// TIA Portal project "Catalyst_syzygy_v2.1" (V17)

(* hardware
DEVICE "S7-1500R/H system_1"  S7-1500R/H-Station
   slot 0: "Rail_0"  Rack  6ES7 590-1***0-0AA0
   slot 1: "Rail_1"  Rack  6ES7 590-1***0-0AA0
   slot 1: "Catalyst_PLC_1"  CPU 1515R-2 PN  6ES7 515-2RM00-0AB0  V2.9
      slot 3: "CPU display_1"  6ES7591-1BA00-0AA0
      slot 32768: "PROFINET interface_1"  X1
         slot 32769: "Port_1"  X1 P1
         slot 32770: "Port_2"  X1 P2
      slot 33024: "PROFINET interface_2"  X2
         slot 33025: "Port_1"  X2 P1
   slot 1: "Catalyst_PLC_2"  CPU 1515R-2 PN  6ES7 515-2RM00-0AB0  V2.9
      slot 3: "CPU display_1"  6ES7591-1BA00-0AA0
      slot 32768: "PROFINET interface_1"  X1
         slot 32769: "Port_1"  X1 P1
         slot 32770: "Port_2"  X1 P2
      slot 33024: "PROFINET interface_2"  X2
         slot 33025: "Port_1"  X2 P1
DEVICE "S7-1500/ET200MP station_1"  S7-1500 station
   slot 0: "Rail_0"  Rack  6ES7 590-1***0-0AA0
   slot 1: "CatalystLocalIO_02"  IM 155-5 PN HF  6ES7 155-5AA00-0AC0  V4.2
   slot 2: "LocalIO_02_AI_01"  AI 8xU/I/RTD/TC ST  6ES7 531-7KF00-0AB0  V2.2
   slot 3: "LocalIO_02_AI_02"  AI 8xU/I/RTD/TC ST  6ES7 531-7KF00-0AB0  V2.2
   slot 4: "LocalIO_02_AI_03"  AI 8xU/I/RTD/TC ST  6ES7 531-7KF00-0AB0  V2.2
   slot 5: "LocalIO_02_AI_04"  AI 8xU/I/RTD/TC ST  6ES7 531-7KF00-0AB0  V2.2
   slot 6: "LocalIO_02_AI_05"  AI 8xU/I/RTD/TC ST  6ES7 531-7KF00-0AB0  V2.2
   slot 7: "LocalIO_02_AI_06"  AI 8xU/I/RTD/TC ST  6ES7 531-7KF00-0AB0  V2.2
   slot 8: "LocalIO_02_AI_07"  AI 8xU/I/RTD/TC ST  6ES7 531-7KF00-0AB0  V2.2
   slot 9: "LocalIO_02_AQ_01"  AQ 8xU/I HS  6ES7 532-5HF00-0AB0  V2.2
   slot 10: "LocalIO_02_AQ_02"  AQ 8xU/I HS  6ES7 532-5HF00-0AB0  V2.1
   slot 11: "LocalIO_02_AQ_03"  AQ 8xU/I HS  6ES7 532-5HF00-0AB0  V2.2
DEVICE "S7-1500/ET200MP station_2"  S7-1500 station
   slot 0: "Rail_0"  Rack  6ES7 590-1***0-0AA0
   slot 1: "CatalystLocalIO_01"  IM 155-5 PN HF  6ES7 155-5AA00-0AC0  V4.4
   slot 2: "LocalIO_01_DI_01"  DI 16x24VDC HF  6ES7 521-1BH00-0AB0  V2.2
   slot 3: "LocalIO_01_DI_02"  DI 16x24VDC HF  6ES7 521-1BH00-0AB0  V2.2
   slot 4: "LocalIO_01_DI_03"  DI 16x24VDC HF  6ES7 521-1BH00-0AB0  V2.2
   slot 5: "LocalIO_01_DI_04"  DI 16x24VDC HF  6ES7 521-1BH00-0AB0  V2.2
   slot 6: "LocalIO_01_DI_05"  DI 16x24VDC HF  6ES7 521-1BH00-0AB0  V2.2
   slot 7: "LocalIO_01_DI_06"  DI 16x24VDC HF  6ES7 521-1BH00-0AB0  V2.2
   slot 8: "LocalIO_01_DQ_01"  DQ 16x24VDC/0.5A HF  6ES7 522-1BH01-0AB0  V1.1
   slot 9: "LocalIO_01_DQ_02"  DQ 16x24VDC/0.5A HF  6ES7 522-1BH01-0AB0  V1.1
   slot 10: "LocalIO_01_DQ_03"  DQ 16x24VDC/0.5A HF  6ES7 522-1BH01-0AB0  V1.1
   slot 11: "LocalIO_01_DQ_04"  DQ 16x24VDC/0.5A HF  6ES7 522-1BH01-0AB0  V1.1
   slot 12: "LocalIO_01_AI_01"  AI 8xU/I/RTD/TC ST  6ES7 531-7KF00-0AB0  V2.2
   slot 13: "LocalIO_01_AI_02"  AI 8xU/I/RTD/TC ST  6ES7 531-7KF00-0AB0  V2.2
   slot 14: "LocalIO_01_AI_03"  AI 8xU/I/RTD/TC ST  6ES7 531-7KF00-0AB0  V2.2
DEVICE "SITOP station_1"  SITOP-Station
   slot 0: "Rack_0"  Rail
   slot 0: "UPS1600"  UPS1600 40A PN  6EP4137-3AB00-2AY0  V2.5
   slot 1: "BAT1600 EX Pb 24V 12Ah_1"  Battery module EX 12Ah Pb  6EP4135-0GL00-0AY0  V1.0
DEVICE "GSD device_1"  GSD.Device.PN
   slot 0: "Rack"  Rack  V1.0
   slot 0: "R-402_DO"  FEN20-4DIP-4DXP  6931090  SW V 1.7.14
      slot 0: "DAP v3.1"  DAP v3.1
      slot 1: "PN-IO"  PN-IO
         slot 1: "Port 1"  Port 1
         slot 2: "Port 2"  Port 2
      slot 1: "4DIP-DXP_1"  4DIP-DXP
         slot 0: "4DIP-DXP"  4DIP-DXP
DEVICE "ET 200SP station_1"  ET 200SP-Station
   slot 0: "Rack_0"  Rack  6ES5 710-8MAx1
   slot 0: "Centrifuge_RIO"  IM 155-6 PN/2 HF  6ES7 155-6AU01-0CN0  V4.2
   slot 1: "DI 8x24VDC ST_1"  DI 8x24VDC ST  6ES7 131-6BF01-0BA0  V0.0
      slot 1: "DI 8x24VDC ST_1"  DI 8x24VDC ST
   slot 2: "DI 8x24VDC ST_2"  DI 8x24VDC ST  6ES7 131-6BF01-0BA0  V0.0
      slot 1: "DI 8x24VDC ST_2"  DI 8x24VDC ST
   slot 3: "DQ 8x24VDC/0.5A ST_1"  DQ 8x24VDC/0.5A ST  6ES7 132-6BF01-0BA0  V0.0
      slot 1: "DQ 8x24VDC/0.5A ST_1"  DQ 8x24VDC/0.5A ST
   slot 4: "AI 4xI 2-,4-wire ST_1"  AI 4xI 2-,4-wire ST  6ES7 134-6GD01-0BA1  V2.0
      slot 1: "AI 4xI 2-,4-wire ST_1"  AI 4xI 2-,4-wire ST
   slot 5: "AQ 4xU/I ST_1"  AQ 4xU/I ST  6ES7 135-6HD00-0BA1  V1.1
      slot 1: "AQ 4xU/I ST_1"  AQ 4xU/I ST
   slot 6: "Server module_1"  Server module  6ES7 193-6PA00-0AA0  V1.1
      slot 1: "Server module_1"  Server module
   slot 127: "BA 2xRJ45"  BA 2xRJ45  6ES7 193-6AR00-0AA0  V0.0
      slot 1: "Port_1"  X1 P1 R  6ES7 193-6AR00-0AA0  V0.0
      slot 2: "Port_2"  X1 P2 R  6ES7 193-6AR00-0AA0  V0.0
DEVICE "GSD device_2"  GSD.Device.PN
   slot 0: "Rack"  Rack  V1.0
   slot 0: "MIXER_T103_VFD"  SINAMICS G120C PN V4.7  6SL3 210-1KExx-xxFx  V4.70
      slot 0: "SINAMICS G120C PN V4.7"  SINAMICS G120C PN V4.7
      slot 1: "PN-IO"  PN-IO
         slot 1: "Port 1"  Port 1
         slot 2: "Port 2"  Port 2
      slot 1: "Drive_1"  Drive
         slot 0: "Module Access Point"  Module Access Point
   slot 2: "Standard telegram 1, PZD-2/2"  Standard telegram 1, PZD-2/2
*)

// ===== PLC "Catalyst_PLC_1"  CPU 1515R-2 PN =====

VAR_GLOBAL   // PLC tag table "Default tag table"
   "Tag_1" AT %T64435 : Timer;
   "Tag_2" AT %T65435 : Timer;
   "moxa_test" AT %M7.2 : Bool;
   "Tag_3" AT %MB3170 : Byte;
   "testdt" AT %MD26 : DInt;
   "addrsscode" AT %MB30 : Byte;
   "addrsscode(1)" AT %MB31 : Byte;
END_VAR

VAR_GLOBAL   // PLC tag table "AQ"
   "ZR-P101A" AT %QW16 : Int;   // P101A discharge pump motor B remote setpoint
   "ZR-P101B" AT %QW18 : Int;   // P101B discharge pump motor B remote setpoint
   "ZR-P102A" AT %QW20 : Int;   // P102A discharge pump motor B remote setpoint
   "ZR-P102B" AT %QW22 : Int;   // P102B discharge pump motor B remote setpoint
   "VFD-T103" AT %QW10 : Int;   // T103 agitator VFD
   "OFF_SQ" AT %M2.1 : Bool;
   "INT_SQ" AT %M2.2 : Bool;
   "ACK_EF" AT %M2.3 : Bool;
   "S_PREV" AT %M2.4 : Bool;
   "S_NEXT" AT %M2.5 : Bool;
   "SW_AUTO" AT %M2.6 : Bool;
   "SW_TAP" AT %M2.0 : Bool;
   "sW_TOP" AT %M2.7 : Bool;
   "SW_MAN" AT %M3.0 : Bool;
   "S_SEL" AT %MW4 : Int;
   "S_ON" AT %M3.1 : Bool;
   "S_OFF" AT %M3.2 : Bool;
   "T_PUSH" AT %M3.3 : Bool;
END_VAR

VAR_GLOBAL   // PLC tag table "ZSO"
   "ZSO-1041" AT %I0.0 : Bool;   // T-101 Water valve open
   "ZSO-1011" AT %I0.3 : Bool;   // T-101 outlet valve open
   "ZSO-1013" AT %I0.5 : Bool;   // T-101 Flow to R-201/202 open
   "ZSO-1042" AT %I0.7 : Bool;   // T-102 Water Valve open
   "ZSO-1021" AT %I1.2 : Bool;   // T-102 Outlet Valve open
   "ZSO-1023" AT %I1.4 : Bool;   // T-102 Flow to R-201/202 open
   "ZSO-1043" AT %I1.6 : Bool;   // R-201 Water Valve open
   "ZSO-1044" AT %I2.0 : Bool;   // R-202 Water Valve open
   "ZSO-2011" AT %I2.2 : Bool;   // T-101 to R-201 Valve open
   "ZSO-2012" AT %I2.4 : Bool;   // T-101 to R-202 Valve open
   "ZSO-2021" AT %I2.6 : Bool;   // T-102 to R-201 Valve open
   "ZSO-2022" AT %I3.0 : Bool;   // T-102 to R-202 Valve open
   "ZSO-2013" AT %I3.3 : Bool;   // R-201 Outlet Valve open
   "ZSO-2023" AT %I3.5 : Bool;   // R-202 Outlet Valve open
   "ZSO-1031" AT %I3.7 : Bool;   // R-201/202 to T-103 Valve open
   "ZSC-1031" AT %I4.0 : Bool;   // R-201/202 to T-103 Valve closed
   "ZSO-1032" AT %I4.2 : Bool;   // T-103 Outlet Valve open
   "ZSO-3011" AT %I4.4 : Bool;   // T-103 to C-301 Valve open
   "ZSO-3012" AT %I4.6 : Bool;   // C-301 Recirc Valve open
   "ZSO-3013" AT %I5.0 : Bool;   // C-301 to ST-301 Valve open
   "ZSO-1045" AT %I5.2 : Bool;   // C-301 Water Valve open
   "ZSO-4011" AT %I5.4 : Bool;   // R-401 Water Trap Valve open
   "ZSO-1033" AT %I7.4 : Bool;   // T-103 Recirc Valve Open
   "ZSO-4024" AT %I8.0 : Bool;   // AIR VALVE OPEN
   "ZSO-4025" AT %I8.2 : Bool;   // N2 VALVE OPEN
END_VAR

VAR_GLOBAL   // PLC tag table "ZSQ"
   "XV-1041" AT %Q1.0 : Bool;   // T-101 Water Valve
   "XV-1011" AT %Q1.1 : Bool;   // T-101 Outlet Valve
   "XV-1021" AT %Q1.3 : Bool;   // T-102 Outlet Valve
   "XV-3011" AT %Q2.6 : Bool;   // T-103 to C-301 Valve
   "XV-3012" AT %Q2.7 : Bool;   // C-301 Recirc Valve
   "XV-1033" AT %Q3.3 : Bool;   // T-103 Recirc Valve
   "XV-4024" AT %Q4.0 : Bool;   // H2 Air Valve
   "XV-1042" AT %Q1.2 : Bool;   // T-102 Water Valve
   "XV-1043" AT %Q1.4 : Bool;   // R-201 Water Valve
   "XV-1044" AT %Q1.5 : Bool;   // R-202 Water Valve
   "XV-2011" AT %Q1.6 : Bool;   // T-101 to R-201 Valve
   "XV-2012" AT %Q1.7 : Bool;   // T-101 to R-202 Valve
   "XV-2021" AT %Q2.0 : Bool;   // T-102 to R-201 Valve
   "XV-2022" AT %Q2.1 : Bool;   // T-102 to R-202 Valve
   "XV-2013" AT %Q2.2 : Bool;   // R-201 Outlet Valve
   "XV-2023" AT %Q2.3 : Bool;   // R-202 Outlet Valve
   "XV-1031" AT %Q2.4 : Bool;   // R-201/202 to T-103 Valve
   "XV-1032" AT %Q2.5 : Bool;   // T-103 Outlet Valve
   "XV-3013" AT %Q3.0 : Bool;   // C-301 Water Valve
   "XV-1045" AT %Q3.1 : Bool;   // C-301 Water Valve
   "XV-4011" AT %Q3.2 : Bool;   // R-401 Water Trap Valve
   "XV-4025" AT %Q4.1 : Bool;   // N2 Air Valve
   "XV-1013" AT %Q4.3 : Bool;   // T-101 Flow to R-201/202
   "XV-1023" AT %Q4.4 : Bool;   // T-102 Flow to R-201/202
END_VAR

VAR_GLOBAL   // PLC tag table "ZSC"
   "ZSC-1041" AT %I0.1 : Bool;   // T-101 Water valve closed
   "ZSC-1011" AT %I0.4 : Bool;   // T-101 outlet valve closed
   "ZSC-1013" AT %I0.6 : Bool;   // T-101 Flow to R-201/202 closed
   "ZSC-1042" AT %I1.0 : Bool;   // T-102 Water Valve closed
   "ZSC-1021" AT %I1.3 : Bool;   // T-102 Outlet Valve closed
   "ZSC-1023" AT %I1.5 : Bool;   // T-102 Flow to R-201/202 closed
   "ZSC-1043" AT %I1.7 : Bool;   // R-201 Water Valve closed
   "ZSC-1044" AT %I2.1 : Bool;   // R-202 Water Valve closed
   "ZSC-2011" AT %I2.3 : Bool;   // T-101 to R-201 Valve closed
   "ZSC-2012" AT %I2.5 : Bool;   // T-101 to R-202 Valve closed
   "ZSC-2021" AT %I2.7 : Bool;   // T-102 to R-201 Valve closed
   "ZSC-2022" AT %I3.1 : Bool;   // T-102 to R-202 Valve closed
   "ZSC-2013" AT %I3.4 : Bool;   // R-201 Outlet Valve closed
   "ZSC-2023" AT %I3.6 : Bool;   // R-202 Outlet Valve closed
   "ZSC-1032" AT %I4.3 : Bool;   // T-103 Outlet Valve closed
   "ZSC-3011" AT %I4.5 : Bool;   // T-103 to C-301 Valve closed
   "ZSC-3012" AT %I4.7 : Bool;   // C-301 Recirc Valve closed
   "ZSC-3013" AT %I5.1 : Bool;   // C-301 to ST-301 Valve closed
   "ZSC-1045" AT %I5.3 : Bool;   // C-301 Water Valve closed
   "ZSC-4011" AT %I5.5 : Bool;   // R-401 Water Trap Valve closed
   "ZSC-1033" AT %I7.5 : Bool;   // T-103 Recirc Valve Closed
   "ZSC-4024" AT %I8.1 : Bool;   // AIR VALVE CLOSED
   "ZSC-4025" AT %I8.3 : Bool;   // N2 VALVE CLOSED
END_VAR

VAR_GLOBAL   // PLC tag table "PH"
   "pH-2021" AT %IW64 : Int;   // R-202 pH #1
   "pH-2022" AT %IW66 : Int;   // R-202 pH #2
   "pH-2011" AT %IW34 : Int;   // R-201 pH #1
   "pH-2012" AT %IW36 : Int;   // R-201 pH #2
END_VAR

VAR_GLOBAL   // PLC tag table "LT"
   "LT-2021" AT %IW68 : Int;   // R-202 Level
   "LT-1031" AT %IW74 : Int;   // T-103 Level
   "LT-2011" AT %IW38 : Int;   // R-201 Level
   "LT-1051" AT %IW122 : Int;   // T-105 LeveL
   "LT-1011" AT %IW16 : Int;   // T-101 LeveL
   "LT-1021" AT %IW26 : Int;   // T-102 LeveL
   "LT-1061" AT %IW140 : Int;   // T-106 Level
END_VAR

VAR_GLOBAL   // PLC tag table "FT"
   "FT-3011" AT %IW80 : Int;   // T-103 to C-301 Flow
   "FT-2022" AT %IW28 : Int;   // T-102 to R-202 Flow
   "FT-1045" AT %IW94 : Int;   // C-301 Water Flow
   "FT-1021" AT %IW48 : Int;   // T-102 Recirc Flow
   "FT-1043" AT %IW50 : Int;   // R-201 Water Flow
   "FT-1044" AT %IW52 : Int;   // R-202 Water Flow
   "FT-2011" AT %IW54 : Int;   // T-101 to R-201 Flow
   "FT-2012" AT %IW56 : Int;   // T-101 to R-202 Flow
   "FT-2021" AT %IW58 : Int;   // T-102 to R-201 Flow
   "FT-3012" AT %IW142 : Int;   // C-301 Outlet Flow
   "FT-1041" AT %IW14 : Int;   // T-101 Water Flow
   "FT-1011" AT %IW22 : Int;   // T-101 Recirc Flow
   "FT-1042" AT %IW24 : Int;   // T-102 Recirc Flow
END_VAR

VAR_GLOBAL   // PLC tag table "AT"
   "AT-3011" AT %IW90 : Int;   // C-301 Nitrates Analyzer
   "AT-3012" AT %IW92 : Int;   // C-301 Turbidity Analyzer
   "AT-4221" AT %IW82 : Int;   // C-402 Calcination O2 Analyzer #1
   "AT-4222" AT %IW84 : Int;   // C-402 Calcination O2 Analyzer #2
END_VAR

VAR_GLOBAL   // PLC tag table "ZT"
   "ZT-T101" AT %IW104 : Int;   // T101 agitator speed
   "ZT-T102" AT %IW106 : Int;   // T102 agitator speed
   "ZT-R201" AT %IW108 : Int;   // R201 agitator speed
   "ZT-R202" AT %IW110 : Int;   // R202 agitator speed
END_VAR

VAR_GLOBAL   // PLC tag table "GD"
   "GD-H2-2" AT %IW120 : Int;   // Hydrogen Gas Detector #2
   "GD-H2-1" AT %IW118 : Int;   // Hydrogen Gas Detector #1
   "GD-CO" AT %IW96 : Int;
END_VAR

VAR_GLOBAL   // PLC tag table "FV"
   "FV-2022" AT %QW64 : Int;
   "FV-2021" AT %QW62 : Int;
   "FV-2012" AT %QW60 : Int;
   "FV-2011" AT %QW58 : Int;
   "FV-3011" AT %QW30 : Int;
   "AN-1000" AT %IW114 : Int;
END_VAR

VAR_GLOBAL   // PLC tag table "VFD"
   "VFD-R202" AT %QW72 : Int;
   "VFD-R201" AT %QW70 : Int;
   "VFD-T102" AT %QW68 : Int;
   "VFD-T101" AT %QW66 : Int;
   "VFD-C301R" AT %QW50 : Int;   // C301 rental centrifuge remote setpoin
END_VAR

VAR_GLOBAL   // PLC tag table "SP"
   "ZR-C301R" AT %I7.0 : Bool;   // C301 rental centrifuge remote setpoint
   "R-401" AT %QW24 : Int;   // R-401 Temp Setpoint
   "TR-H201" AT %QW28 : Int;   // H-201 Temperature Control Output
END_VAR

VAR_GLOBAL   // PLC tag table "Enable PMP"
   "HS-P201A" AT %Q5.0 : Bool;   // P201A discharge pump motor A - Enable
   "HS-P201B" AT %Q5.1 : Bool;   // P201B discharge pump motor B - Enable
   "HS-P202A" AT %Q5.4 : Bool;   // P202A discharge pump motor A - Enable
   "HS-P202B" AT %Q5.5 : Bool;   // P202B discharge pump motor B - Enable
   "HS-P103A" AT %Q6.0 : Bool;   // P103A discharge pump motor A - Enable
   "HS-P103B" AT %Q6.1 : Bool;   // P103B discharge pump motor B - Enable
   "HR-T101" AT %Q3.4 : Bool;   // T101 agitator motor - Enable
   "HR-T102" AT %Q3.5 : Bool;   // T102 agitator motor - Enable
   "HR-R201" AT %Q3.6 : Bool;   // R201 agitator motor - Enable
   "HR-R202" AT %Q3.7 : Bool;   // R202 agitator motor - Enable
   "HS-P101A" AT %Q7.2 : Bool;   // P101A discharge pump motor A - Enable
   "HS-P101B" AT %Q7.3 : Bool;   // P101B discharge pump motor B - Enable
   "HS-P102A" AT %Q7.4 : Bool;   // P102A discharge pump motor A - Enable
   "HS-P102B" AT %Q7.5 : Bool;   // P102B discharge pump motor B - Enable
   "H-201" AT %Q0.1 : Bool;   // H-201 (Future)
END_VAR

VAR_GLOBAL   // PLC tag table " Start Remote"
   "HS-C301" AT %Q6.2 : Bool;   // C301 centirfuge motor - Start remote
   "HS-C301A" AT %Q6.3 : Bool;   // P301A discharge pump motor A - Start Remote
   "HS-C301B" AT %Q6.4 : Bool;   // P301B discharge pump motor B - start remote
   "HS-P104C" AT %Q6.5 : Bool;   // P104C discharge pump motor C - Start Remote
   "HS-P104A" AT %Q6.6 : Bool;   // P104A discharge pump motor A - Start Remote
   "HS-P104B" AT %Q6.7 : Bool;   // P104B discharge pump motor B - Start Remote
END_VAR

VAR_GLOBAL   // PLC tag table "POWER_SUPPLY"
   "SP1-11" AT %I8.4 : Bool;
   "SP2-11" AT %I8.5 : Bool;
   "SP1-13" AT %I8.6 : Bool;
   "SP2-13" AT %I8.7 : Bool;
   "MFC-4011-F" AT %MW8 : Int;
   "MFC-4024-F" AT %MW12 : Int;
   "MFC-4025-F" AT %MW14 : Int;
   "MFC-4011-P" AT %MW10 : Int;
   "MFC-4024-P" AT %MW16 : Int;
END_VAR

VAR_GLOBAL   // PLC tag table "agitator motor running"
   "ZR-T101" AT %I5.6 : Bool;   // T101 agitator motor running
   "ZR-T102" AT %I6.0 : Bool;   // T102 agitator motor running
   "ZR-R201" AT %I6.2 : Bool;   // R201 agitator motor running
   "ZR-R202" AT %I6.4 : Bool;   // R202 agitator motor running
END_VAR

VAR_GLOBAL   // PLC tag table " agitator motor - Hand switch Local"
   "HS-T101L" AT %I5.7 : Bool;   // T101 agitator motor - Hand switch Local
   "HS-T102L" AT %I6.1 : Bool;   // T102 agitator motor - Hand switch Local
   "HS-R201L" AT %I6.3 : Bool;   // R201 agitator motor - Hand switch Local
   "HS-R202L" AT %I6.5 : Bool;   // R202 agitator motor - Hand switch Local
   "OFF_SQ_1" AT %M3.4 : Bool;
   "INT_SQ_1" AT %M3.5 : Bool;
   "INT_SQ_2" AT %M3.6 : Bool;
   "OFF_SQ_2" AT %M3.7 : Bool;
   "rst" AT %M6.3 : Bool;
   "TEST_BIT" AT %M6.4 : Bool;
   "MFC-4025-P" AT %MW18 : Int;
   "MFC-4011-T" AT %MW20 : Int;
   "MFC-4024-T" AT %MW22 : Int;
   "MFC-4025-T" AT %MW24 : Int;
   "testTimerCalcination" AT %M7.1 : Bool;
   "TE-402A_Sim" AT %MW32 : Int;
   "TE-402B_Sim" AT %MW34 : Int;
END_VAR

VAR_GLOBAL   // PLC tag table "LSHH"
   "LSHH-1011" AT %I0.2 : Bool;   // T-101 High High Level Switch
   "LSHH-1021" AT %I1.1 : Bool;   // T-102 High High Level Switch
   "LSHH-2011" AT %I3.2 : Bool;   // R-201 High High Level Switch
   "LSHH-1031" AT %I4.1 : Bool;   // T-103 High High Level Switch
   "LSHH-2021" AT %I7.3 : Bool;   // R-202 High High Level Switch
   "LSHH-1051" AT %I7.6 : Bool;   // T-105 High High Level Switch
END_VAR

VAR_GLOBAL   // PLC tag table "PT"
   "PT-202A" AT %IW12 : Int;   // P-202A Pressure
   "PT-103B" AT %IW78 : Int;   // P-103B Pressure
   "PT-301A" AT %IW86 : Int;   // P-301A Pressure
   "PT-301B" AT %IW88 : Int;   // P-301B Pressure
   "PT-104A" AT %IW148 : Int;   // PT-104A
   "PT-104B" AT %IW150 : Int;   // PT-104B
   "PT-202B" AT %IW70 : Int;   // P-202B Pressure
   "PT-101A" AT %IW18 : Int;   // P-101A Dischare Pressure
   "PT-101B" AT %IW20 : Int;   // P-101B Discharge Pressure
   "PT-102A" AT %IW44 : Int;   // P-102A Dischare Pressure
   "PT-102B" AT %IW46 : Int;   // P-102B Discharge Pressure
   "PT-201A" AT %IW40 : Int;   // P-201A Pressure
   "PT-201B" AT %IW42 : Int;   // P-201B Pressure
   "PT-103A" AT %IW76 : Int;   // P-103A Pressure
END_VAR

VAR_GLOBAL   // PLC tag table "TT"
   "TT-2021" AT %IW60 : Int;   // R-202 Temperature #1
   "TT-2022" AT %IW62 : Int;   // R-202 Temperature #2
   "TT-1031" AT %IW72 : Int;   // T-103 Temperature
   "TE-401A" AT %IW132 : Int;   // R-401 Temperature #1
   "TE-401B" AT %IW134 : Int;   // R-401 Temperature #2
   "TE-401C" AT %IW136 : Int;   // R-401 Temperature #3
   "TT-2011" AT %IW30 : Int;   // R-201 Temperature #1
   "TT-2012" AT %IW32 : Int;   // R-201 Temperature #2
   "ENC_RTD_PT-100" AT %IW126 : Int;   // Enclosure RTD PT-100
   "TE-H201" AT %IW112 : Int;   // H-201 Temperature
   "TE-402A" AT %IW156 : Int;   // R-402 Temperature #1
   "TE-402B" AT %IW158 : Int;   // R-402 Temperature #2
   "TE-402C" AT %IW160 : Int;   // R-402 Temperature #3
   "TE-402D" AT %IW162 : Int;   // R-402 Temperature #4
   "TE-401D" AT %IW138 : Int;   // R-401 Temperature #4
   "TE-402E" AT %IW164 : Int;   // R-402 Temperature #5
END_VAR

VAR_GLOBAL CONSTANT   // PLC tag table "StateMachineConts"
   "T-101HighLimit" : Real := 75.00;   // This Value is a Percentage of the Tank
   "T-101HighHighLimit" : Real := 80.00;   // This Value is a Percentage of the Tank
   "Pumps101TramisttersHighLimit" : Real := 126.00;   // This Value is in PSI
   "Pumps101TramisttersHighHighLimit" : Real := 129.00;   // This Value is IN PSI
   "T-102HighLimit" : Real := 75.00;   // This Value is a Percentage of the Tank
   "T-102HighHighLimit" : Real := 80.00;   // This Value is a Percentage of the Tank
   "Pumps102TramisttersHighLimit" : Real := 126.00;   // This Value is in PSI
   "Pumps102TramisttersHighHighLimit" : Real := 129.00;   // This Value is IN PSI
   "SingleReactorMaxLevelBatchSize" : Real := 160.00;
   "ReactorMinLevelBatchSize" : Real := 40.00;
   "ReactorLowLevelSetpoint" : Real := 2.0;   // This Value is a Percentage of the Tank
   "WashLowLevelSetpoint" : Real := 2.0;   // This is scale in Percentage
   "MixLowLevelSetpoint" : Real := 2.0;   // This Value is a Percentage of the Tank
   "MinimunFlowForTotalizers" : Real := 0.01;
   "ReactorVFDSpeed" : Real := 65.00;   // Percentannce Value 0-100%
   "MixTanksVFDSpeedSetpointLow" : Real := 70.0;   // Percentannce Value 0-100%
   "MixTanksVFDSpeedSetpointHigh" : Real := 80.0;   // Percentannce Value 0-100%
   "ReactorBatchTemp" : Real := 40.00;
   "VFDminimunReadSpeedFilter" : Int := 38;
   "SoluctionTanksLowSpeedMaxvalue" : Real := 20.5;
   "SoluctionTanksHighSpeedMinValue" : Real := 20.6;
   "AnalyzerLowLevelSetpoint" : Real := 5.0;   // Analyzer TX Minimun Value
   "CoolingLowLevelSetpoint" : Real := 2.0;   // This Value is a Percentage of the Tank
   "ReactorLowExitPressurelSetpoint" : Real := 0.5;   // PSI
   "CentrifugeSpeed" : Real := 500.0;
END_VAR

VAR_GLOBAL   // PLC tag table "Memory_data"
   "Clock_0.5Hz" AT %M0.7 : Bool;
   "AlwaysTRUE" AT %M1.2 : Bool;
   "DiagStatusUpdate" AT %M1.1 : Bool;
   "AlwaysFALSE" AT %M1.3 : Bool;
   "Clock_1Hz" AT %M0.5 : Bool;
   "Clock_10Hz" AT %M0.0 : Bool;
   "Clock_Byte" AT %MB0 : Byte;
   "Clock_1.25Hz" AT %M0.4 : Bool;
   "Clock_2Hz" AT %M0.3 : Bool;
   "FirstScan" AT %M1.0 : Bool;
   "System_Byte" AT %MB1 : Byte;
   "Clock_5Hz" AT %M0.1 : Bool;
   "Clock_0.625Hz" AT %M0.6 : Bool;
   "Clock_2.5Hz" AT %M0.2 : Bool;
   "BYPASS_1" AT %M6.5 : Bool;
   "BYPASS_2" AT %M6.6 : Bool;
   "BYPASS_3" AT %M6.7 : Bool;
   "BYPASS_4" AT %M7.0 : Bool;
   "BYPASS" AT %M6.0 : Bool;
   "bit2" AT %M6.2 : Bool;
   "bit" AT %M6.1 : Bool;
END_VAR

VAR_GLOBAL   // PLC tag table "Centrifuge_IO"
   "CentrifugeVibrationFault" AT %I190.0 : Bool;   // (VTM-8) Vibration Fault on Centrifuge
   "E-STOP_FromCentrifuge" AT %I190.1 : Bool;   // E-STOP from Centrifuge
   "CentrifugeSystemFault" AT %I190.2 : Bool;   // Centrifuge System Fault
   "CentrifugeBasketFull" AT %I190.3 : Bool;   // Centrifuge Basket Full
   "CentrifugeCoverLocked" AT %I190.4 : Bool;   // Centrifuge Cover Locked 1 = Locked, 0= Unlocked
   "CentrifugeFeelerRetracted" AT %I190.5 : Bool;   // Centrifuge Feeler Retracted
   "Tag_7" AT %I190.6 : Bool;
   "Tag_8" AT %I190.7 : Bool;
   "CentrifugeStartCmd" AT %Q9.0 : Bool;   // Centrifuge Start Command
   "E-STOP_ToCentrifuge" AT %Q9.1 : Bool;   // E-STOP to Centrifuge from PLC. 1=OK
   "RetFeelerAndFaultReset" AT %Q9.2 : Bool;   // Retrac Feeler and Fault Reset
   "FeelerEngage" AT %Q9.3 : Bool;   // Feeler Engage
   "CentrifugeStopCmd" AT %Q9.4 : Bool;   // Centrifuge Stop Command
   "Tag_6" AT %Q9.5 : Bool;
   "Tag_7(1)" AT %Q9.6 : Bool;
   "Tag_8(1)" AT %Q9.7 : Bool;
   "CentrifugeVibrationTransmitter" AT %IW182 : Int;   // Centrifuge Vibration Transmitter
   "CentrifugeActualSpeed" AT %IW184 : Int;   // Centrifuge Actual Speed Feedback
   "Tag_3(1)" AT %IW186 : Int;
   "Tag_4" AT %IW188 : Int;
END_VAR

VAR_GLOBAL CONSTANT   // PLC tag table "ModbusIDs"
   "MFC-4011_MBID" : Conn_Any := 1;
   "MFC-4012_MBID" : Conn_Any := 2;
   "MFC-4021_MBID" : Conn_Any := 33;
   "MFC-4024_MBID" : Conn_Any := 34;
   "TC-4011A_MBID" : Conn_Any := 30;
   "TC-4011B_MBID" : Conn_Any := 31;
   "TC-4011C_MBID" : Conn_Any := 32;
   "pH-2011_12_MBID" : Conn_Any := 3;
   "pH-2021_22_MBID" : Conn_Any := 4;
   "Analizer_R-401_MBID" : Conn_Any := 35;
END_VAR

TYPE "ModBus_Data"
   STRUCT
      Slaves : Struct
         Slave1 : Array[1..12] of Int;
         Slave2 : Array[1..12] of Int;
         Slave3 : Array[1..12] of Int;
      END_STRUCT;
   END_STRUCT;
END_TYPE

TYPE "EurothermCtls_UDT"
   STRUCT
      Read : Struct
         WorkingSP : Real;   // Running Setpoints (From Controller)
         PV : Real;   // Process Value (From Controller)
         OP : Real;   // Controller Output (From Controller)
         FaultTemperature : Bool;
      END_STRUCT;
      Write : Struct
         Dwell : Int;   // Dwell Duration in Hours
         CMD : Int;   // 0= Stop, 1=Run
         SP : Real;   // SetPoint (To controller)
         RampSp : Int;   // Ramp SP Degree per min
      END_STRUCT;
   END_STRUCT;
END_TYPE

TYPE "AlicatCtl_UDT"
   STRUCT
      CMD_ID : Int;   // Command ID (See Modbus RTU Manual)
      CMD_Arg : Int;   // Command Argument (See Modbus RTU Manual)
      SP : Real;   // Flow SP sent to the Flow Controller
      PV : Real;   // Flow Process Value Controlled
      Status : Struct
         Fbk : Real;   // Feedback of the Control Valve Position
         CommFault : Bool;
      END_STRUCT;
   END_STRUCT;
END_TYPE

TYPE "ModBus_DataP"
   STRUCT
      Slaves : Struct
         Data : Array[1..3, 1..12] of Int;
      END_STRUCT;
   END_STRUCT;
END_TYPE

// folder: Actuator

TYPE "Cmd"
   STRUCT
      Enable : Bool;
      CmdOn : Bool;
      TurningOff : Bool;
      TurningOn : Bool;
   END_STRUCT;
END_TYPE

TYPE "Cmd_VFD"
   STRUCT
      Enable : Bool;   // Enable
      CmdOn : Bool;   // On Command
      Reset : Bool;   // Reset Alarms
      Running : Bool;
      Error : Bool;
      Status : Word;
      TurningOff : Bool;
      TurningOn : Bool;
      p2000 : Real;   // Value from p2000 at VFD Configuration (Starter)
      SP : Real;   // SetPoint (%)
      Fbk : Real;   // Feedback (RPM)
   END_STRUCT;
END_TYPE

TYPE "TC_Read"
   STRUCT
      ActSP : Real;
      PV : Real;
      OP : Real;
      FaultTemperature : Bool;
   END_STRUCT;
END_TYPE

TYPE "TC_Write"
   STRUCT
      Dwell : Int;
      CMD : Int;
      SP : Real;
      RampSp : Int;
   END_STRUCT;
END_TYPE

TYPE "Centrifuge"
   STRUCT
      Enable : Bool;   // Enable
      Start : Bool;   // On Command
      Stop : Bool;
      RetracReset : Bool;
      FeelerEngage : Bool;
      SP : Real;   // SetPoint (%)
      Fbk : Real;   // Feedback (RPM)
   END_STRUCT;
END_TYPE

// folder: HMI

TYPE "ToHMI"
   STRUCT
      EnStopButton : Bool;   // Enable HMI Stop Button
      EnStartButton : Bool;   // Enable HMI Start Button
      EnRestartButton : Bool;
      EnPauseButton : Bool;
      EnOpeRequest : Bool;   // Enable HMI Operator Request Button
      EnEditorButton : Bool;   // Enable HMI Editor Burron Button
      InterlockActivated : Bool;
      Spare01 : Bool;
      Spare02 : Bool;
   END_STRUCT;
END_TYPE

TYPE "FromHMI"
   STRUCT
      Start : Bool;   // Start Sequence
      Stop : Bool;   // Stop Sequence
      Pause : Bool;
      Restart : Bool;
      Initialize : Bool;   // Initialize Sequence
      TankWash : Bool;   // Tank Wash Procedure
      TubeWash : Bool;   // Line Wash Procedure
      Transfer : Bool;
      Receive : Bool;
      Mix : Bool;   // Transfer to Cooling Tank (T-103)
      Pouring : Bool;
      Centrifuge : Bool;   // Transfer to Cooling Tank (T-103)
      Spare01 : Bool;
      Spare02 : Bool;
      Procedure : Int;   // Recipe Procedure
   END_STRUCT;
END_TYPE

// folder: Unit

TYPE "UnitCmds"
   STRUCT
      Start : Bool;
      Hold : Bool;
      Resume : Bool;
      Initialize : Bool;
      TankWash : Bool;
      TubeWash : Bool;
      Transfer : Bool;
      Receive : Bool;
      Mix : Bool;
      Pouring : Bool;
      Centrifuge : Bool;
      Calcination : Bool;   // Calcination Process
      Passivation : Bool;   // Passivation Process
      Reduction : Bool;   // Reduction Process
      ControlledShutdown : Bool;   // Controlled Shurdown command
      Abort : Bool;   // Abort Command
      PermCond : Bool;   // Permanent Condition to Transitions
      IL : Bool;   // IL=1 (Interlocks Good) , IL=0 ESD Activated
      Procedure : Int := 1;   // Recipe Procedure
   END_STRUCT;
END_TYPE

// folder: (top level)

DATA_BLOCK "test_db"   // DB26
{ S7_Optimized_Access := 'TRUE' }
VERSION : 0.1
// stored: InstanceOfName PID_TIA
"PID_TIA"
BEGIN
END_DATA_BLOCK

// folder: Analogs inputs/Trasmitters/Analyzer Trasmitters/Datablocks

DATA_BLOCK "AT-3011_DB"   // DB66
{ S7_Optimized_Access := 'TRUE' }
VERSION : 1.0
// stored: InstanceOfName TX-AI
"TX-AI"
BEGIN
END_DATA_BLOCK

DATA_BLOCK "AT-3012_DB"   // DB67
{ S7_Optimized_Access := 'TRUE' }
VERSION : 1.0
// stored: InstanceOfName TX-AI
"TX-AI"
BEGIN
END_DATA_BLOCK

DATA_BLOCK "AT-4021_DB"   // DB127
{ S7_Optimized_Access := 'TRUE' }
VERSION : 1.0
// stored: InstanceOfName TX-AI
"TX-AI"
BEGIN
   Retain.HMI.Config.ESMXV := 25.0;
END_DATA_BLOCK

DATA_BLOCK "AT-4022_DB"   // DB203
{ S7_Optimized_Access := 'TRUE' }
VERSION : 1.0
// stored: InstanceOfName TX-AI
"TX-AI"
BEGIN
   Retain.HMI.Config.ESMXV := 25.0;
END_DATA_BLOCK

// folder: Analogs inputs/Trasmitters/Flow Trasmitters/Datablocks

DATA_BLOCK "FT-1041_DB"   // DB30
{ S7_Optimized_Access := 'TRUE' }
VERSION : 1.0
// stored: InstanceOfName TX-AI
"TX-AI"
BEGIN
   Retain.HMI.Config.ESMXV := 50.0;
   Retain.HMI.Config.SP.Limits.HH := 45.0;
   Retain.HMI.Config.SP.Limits.H := 40.0;
   Retain.HMI.Config.SP.Limits.L := 5.0;
   Retain.HMI.Config.PT.DBNC.AL := t#20s;
END_DATA_BLOCK

DATA_BLOCK "FT-1011_DB"   // DB33
{ S7_Optimized_Access := 'TRUE' }
VERSION : 1.0
// stored: InstanceOfName TX-AI
"TX-AI"
BEGIN
   Retain.HMI.Config.ESMXV := 10.0;
   Retain.HMI.Config.SP.Limits.HH := 9.0;
   Retain.HMI.Config.SP.Limits.H := 8.0;
END_DATA_BLOCK

DATA_BLOCK "FT-1042_DB"   // DB34
{ S7_Optimized_Access := 'TRUE' }
VERSION : 1.0
// stored: InstanceOfName TX-AI
"TX-AI"
BEGIN
   Retain.HMI.Config.ESMXV := 50.0;
   Retain.HMI.Config.SP.Limits.HH := 45.0;
   Retain.HMI.Config.SP.Limits.H := 40.0;
   Retain.HMI.Config.SP.Limits.L := 5.0;
   Retain.HMI.Config.PT.DBNC.AL := t#20s;
END_DATA_BLOCK

DATA_BLOCK "FT-1021_DB"   // DB38
{ S7_Optimized_Access := 'TRUE' }
VERSION : 1.0
// stored: InstanceOfName TX-AI
"TX-AI"
BEGIN
   Retain.HMI.Config.ESMXV := 10.0;
   Retain.HMI.Config.SP.Limits.HH := 9.0;
   Retain.HMI.Config.SP.Limits.H := 8.0;
END_DATA_BLOCK

DATA_BLOCK "FT-1043_DB"   // DB39
{ S7_Optimized_Access := 'TRUE' }
VERSION : 1.0
// stored: InstanceOfName TX-AI
"TX-AI"
BEGIN
   Retain.HMI.Config.ESMXV := 50.0;
   Retain.HMI.Config.SP.Limits.HH := 45.0;
   Retain.HMI.Config.SP.Limits.H := 40.0;
   Retain.HMI.Config.SP.Limits.L := 5.0;
   Retain.HMI.Config.PT.DBNC.AL := t#20s;
END_DATA_BLOCK

DATA_BLOCK "FT-2011_DB"   // DB40
{ S7_Optimized_Access := 'TRUE' }
VERSION : 1.0
// stored: InstanceOfName TX-AI
"TX-AI"
BEGIN
   Retain.HMI.Config.ESMXV := 5.0;
   Retain.HMI.Config.SP.Limits.HH := 9.0;
   Retain.HMI.Config.SP.Limits.H := 8.0;
END_DATA_BLOCK

DATA_BLOCK "FT-2021_DB"   // DB41
{ S7_Optimized_Access := 'TRUE' }
VERSION : 1.0
// stored: InstanceOfName TX-AI
"TX-AI"
BEGIN
   Retain.HMI.Config.ESMXV := 5.0;
   Retain.HMI.Config.SP.Limits.HH := 9.0;
   Retain.HMI.Config.SP.Limits.H := 8.0;
END_DATA_BLOCK

DATA_BLOCK "FT-2012_DB"   // DB42
{ S7_Optimized_Access := 'TRUE' }
VERSION : 1.0
// stored: InstanceOfName TX-AI
"TX-AI"
BEGIN
   Retain.HMI.Config.ESMXV := 5.0;
   Retain.HMI.Config.SP.Limits.HH := 9.0;
   Retain.HMI.Config.SP.Limits.H := 8.0;
END_DATA_BLOCK

DATA_BLOCK "FT-2022_DB"   // DB43
{ S7_Optimized_Access := 'TRUE' }
VERSION : 1.0
// stored: InstanceOfName TX-AI
"TX-AI"
BEGIN
   Retain.HMI.Config.ESMXV := 5.0;
   Retain.HMI.Config.SP.Limits.HH := 9.0;
   Retain.HMI.Config.SP.Limits.H := 8.0;
END_DATA_BLOCK

DATA_BLOCK "FT-1044_DB"   // DB48
{ S7_Optimized_Access := 'TRUE' }
VERSION : 1.0
// stored: InstanceOfName TX-AI
"TX-AI"
BEGIN
   Retain.HMI.Config.ESMXV := 50.0;
   Retain.HMI.Config.SP.Limits.HH := 45.0;
   Retain.HMI.Config.SP.Limits.H := 40.0;
   Retain.HMI.Config.SP.Limits.L := 5.0;
   Retain.HMI.Config.PT.DBNC.AL := t#20s;
END_DATA_BLOCK

DATA_BLOCK "FT-3011_DB"   // DB63
{ S7_Optimized_Access := 'TRUE' }
VERSION : 1.0
// stored: InstanceOfName TX-AI
"TX-AI"
BEGIN
   Retain.HMI.Config.ESMXV := 5.0;
   Retain.HMI.Config.SP.Limits.HH := 4.5;
   Retain.HMI.Config.SP.Limits.H := 4.0;
   Retain.HMI.Config.PT.DBNC.AL := t#1m;
END_DATA_BLOCK

DATA_BLOCK "FT-1045_DB"   // DB68
{ S7_Optimized_Access := 'TRUE' }
VERSION : 1.0
// stored: InstanceOfName TX-AI
"TX-AI"
BEGIN
   Retain.HMI.Config.ESMXV := 50.0;
   Retain.HMI.Config.SP.Limits.HH := 45.0;
   Retain.HMI.Config.SP.Limits.H := 40.0;
   Retain.HMI.Config.SP.Limits.L := 5.0;
   Retain.HMI.Config.PT.DBNC.AL := t#20s;
END_DATA_BLOCK

DATA_BLOCK "FT-3012_DB"   // DB126
{ S7_Optimized_Access := 'TRUE' }
VERSION : 1.0
// stored: InstanceOfName TX-AI
"TX-AI"
BEGIN
   Retain.HMI.Config.ESMXV := 30.0;
   Retain.HMI.Config.SP.Limits.HH := 28.0;
   Retain.HMI.Config.SP.Limits.H := 25.0;
   Retain.HMI.Config.SP.Limits.L := 2.0;
   Retain.HMI.Config.PT.DBNC.AL := t#30s;
END_DATA_BLOCK

DATA_BLOCK "MFC-4011-F_DB"   // DB161
{ S7_Optimized_Access := 'TRUE' }
VERSION : 1.0
// stored: InstanceOfName TX-AI
"TX-AI"
BEGIN
END_DATA_BLOCK

DATA_BLOCK "MFC-4012-F_DB"   // DB199
{ S7_Optimized_Access := 'TRUE' }
VERSION : 1.0
// stored: InstanceOfName TX-AI
"TX-AI"
BEGIN
END_DATA_BLOCK

DATA_BLOCK "MFC-4024-F_DB"   // DB212
{ S7_Optimized_Access := 'TRUE' }
VERSION : 1.0
// stored: InstanceOfName TX-AI
"TX-AI"
BEGIN
END_DATA_BLOCK

DATA_BLOCK "MFC-4025-F_DB"   // DB215
{ S7_Optimized_Access := 'TRUE' }
VERSION : 1.0
// stored: InstanceOfName TX-AI
"TX-AI"
BEGIN
END_DATA_BLOCK

DATA_BLOCK "AN-1000_DB"   // DB227
{ S7_Optimized_Access := 'TRUE' }
VERSION : 1.0
// stored: InstanceOfName TX-AI
"TX-AI"
BEGIN
END_DATA_BLOCK

DATA_BLOCK "MFC-4021-F_DB"   // DB436
{ S7_Optimized_Access := 'TRUE' }
VERSION : 1.0
// stored: InstanceOfName TX-AI
"TX-AI"
BEGIN
END_DATA_BLOCK

// folder: Analogs inputs/Trasmitters/Hydrogen Gas Trasmitters/Datablocks

DATA_BLOCK "GD-H2-2_DB"   // DB122
{ S7_Optimized_Access := 'TRUE' }
VERSION : 1.0
// stored: InstanceOfName TX-AI
"TX-AI"
BEGIN
END_DATA_BLOCK

DATA_BLOCK "GD-H2-1_DB"   // DB123
{ S7_Optimized_Access := 'TRUE' }
VERSION : 1.0
// stored: InstanceOfName TX-AI
"TX-AI"
BEGIN
END_DATA_BLOCK

DATA_BLOCK "GD-CO_DB"   // DB204
{ S7_Optimized_Access := 'TRUE' }